REGION Network 65: SOLICITAÇÃO DE DESLIGAMENTO DO GRUPO 1
   RUNG wire#powerrail
      Contact( #AUX05 )
      wire#w1
      Contact( #LG1 )
      Contact( #G1L )
      Coil( #SDESG1 )
      wire#w2
      R_Coil( #LG1 )
   END_RUNG
   RUNG wire#powerrail
      Contact( #RTEOKG1 )
      Contact( #G1P )
   END_RUNG wire#w1
   RUNG wire#powerrail
      I_Contact( #G1OK )
   END_RUNG wire#w2
   RUNG wire#powerrail
      Contact( "AlwaysFALSE" )
      { S7_Templates := "SrcType := Int" } EQ_Contact(in1 := #NGS, in2 := 1)
      I_Contact( #G1P )
   END_RUNG wire#w2
   RUNG wire#powerrail
      Contact( "AlwaysFALSE" )
      { S7_Templates := "SrcType := Int" } EQ_Contact(in1 := #NGS, in2 := 2)
      I_Contact( #G1P )
      I_Contact( #G1C1 )
   END_RUNG wire#w2
   RUNG wire#powerrail
      Contact( "AlwaysFALSE" )
      { S7_Templates := "SrcType := Int" } EQ_Contact(in1 := #NGS, in2 := 3)
      I_Contact( #G1P )
      I_Contact( #G1C1 )
      I_Contact( #G1C2 )
   END_RUNG wire#w2
   RUNG wire#powerrail
      Contact( "AlwaysFALSE" )
      { S7_Templates := "SrcType := Int" } EQ_Contact(in1 := #NGS, in2 := 4)
      I_Contact( #G1P )
      I_Contact( #G1C1 )
      I_Contact( #G1C2 )
      I_Contact( #G1C3 )
   END_RUNG wire#w2
   // the same network as SCL:
   #SDESG1 := (#AUX05 OR (#RTEOKG1 AND #G1P)) AND #LG1 AND #G1L;
   IF #SDESG1 OR NOT #G1OK OR ("AlwaysFALSE" AND (#NGS = 1) AND NOT #G1P) OR ("AlwaysFALSE" AND (#NGS = 2) AND NOT #G1P AND NOT #G1C1) OR ("AlwaysFALSE" AND (#NGS = 3) AND NOT #G1P AND NOT #G1C1 AND NOT #G1C2) OR ("AlwaysFALSE" AND (#NGS = 4) AND NOT #G1P AND NOT #G1C1 AND NOT #G1C2 AND NOT #G1C3) THEN
       #LG1 := FALSE;
   END_IF;
END_REGION

REGION Network 66: SOLICITAÇÃO DE DESLIGAMENTO DO GRUPO 2
   #TSDG2(IN := (#SO_D OR NOT #DESAB) AND #G2P, PT := T#5S, ET => #ETTSDG2);   // TON
   #AUX06 := #TSDG2.Q;
END_REGION

REGION Network 67: SOLICITAÇÃO DE DESLIGAMENTO DO GRUPO 2
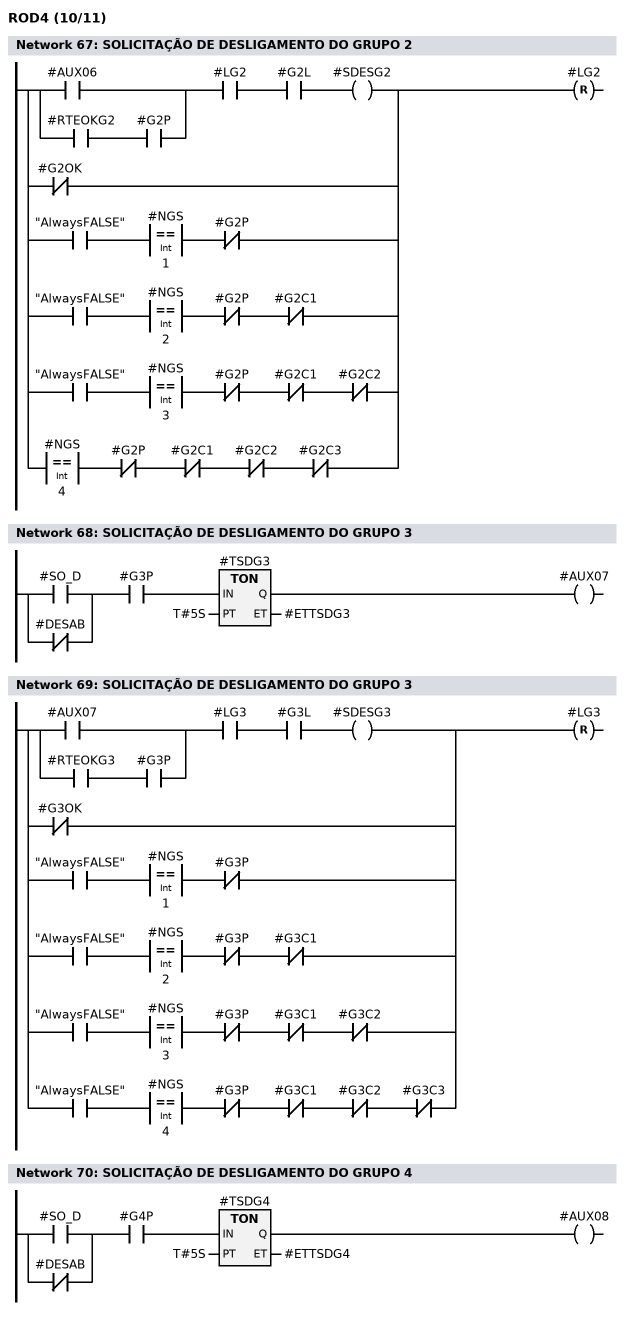
   RUNG wire#powerrail
      Contact( #AUX06 )
      wire#w1
      Contact( #LG2 )
      Contact( #G2L )
      Coil( #SDESG2 )
      wire#w2
      R_Coil( #LG2 )
   END_RUNG
   RUNG wire#powerrail
      Contact( #RTEOKG2 )
      Contact( #G2P )
   END_RUNG wire#w1
   RUNG wire#powerrail
      I_Contact( #G2OK )
   END_RUNG wire#w2
   RUNG wire#powerrail
      Contact( "AlwaysFALSE" )
      { S7_Templates := "SrcType := Int" } EQ_Contact(in1 := #NGS, in2 := 1)
      I_Contact( #G2P )
   END_RUNG wire#w2
   RUNG wire#powerrail
      Contact( "AlwaysFALSE" )
      { S7_Templates := "SrcType := Int" } EQ_Contact(in1 := #NGS, in2 := 2)
      I_Contact( #G2P )
      I_Contact( #G2C1 )
   END_RUNG wire#w2
   RUNG wire#powerrail
      Contact( "AlwaysFALSE" )
      { S7_Templates := "SrcType := Int" } EQ_Contact(in1 := #NGS, in2 := 3)
      I_Contact( #G2P )
      I_Contact( #G2C1 )
      I_Contact( #G2C2 )
   END_RUNG wire#w2
   RUNG wire#powerrail
      { S7_Templates := "SrcType := Int" } EQ_Contact(in1 := #NGS, in2 := 4)
      I_Contact( #G2P )
      I_Contact( #G2C1 )
      I_Contact( #G2C2 )
      I_Contact( #G2C3 )
   END_RUNG wire#w2
   // the same network as SCL:
   #SDESG2 := (#AUX06 OR (#RTEOKG2 AND #G2P)) AND #LG2 AND #G2L;
   IF #SDESG2 OR NOT #G2OK OR ("AlwaysFALSE" AND (#NGS = 1) AND NOT #G2P) OR ("AlwaysFALSE" AND (#NGS = 2) AND NOT #G2P AND NOT #G2C1) OR ("AlwaysFALSE" AND (#NGS = 3) AND NOT #G2P AND NOT #G2C1 AND NOT #G2C2) OR ((#NGS = 4) AND NOT #G2P AND NOT #G2C1 AND NOT #G2C2 AND NOT #G2C3) THEN
       #LG2 := FALSE;
   END_IF;
END_REGION

REGION Network 68: SOLICITAÇÃO DE DESLIGAMENTO DO GRUPO 3
   #TSDG3(IN := (#SO_D OR NOT #DESAB) AND #G3P, PT := T#5S, ET => #ETTSDG3);   // TON
   #AUX07 := #TSDG3.Q;
END_REGION

REGION Network 69: SOLICITAÇÃO DE DESLIGAMENTO DO GRUPO 3
   RUNG wire#powerrail
      Contact( #AUX07 )
      wire#w1
      Contact( #LG3 )
      Contact( #G3L )
      Coil( #SDESG3 )
      wire#w2
      R_Coil( #LG3 )
   END_RUNG
   RUNG wire#powerrail
      Contact( #RTEOKG3 )
      Contact( #G3P )
   END_RUNG wire#w1
   RUNG wire#powerrail
      I_Contact( #G3OK )
   END_RUNG wire#w2
   RUNG wire#powerrail
      Contact( "AlwaysFALSE" )
      { S7_Templates := "SrcType := Int" } EQ_Contact(in1 := #NGS, in2 := 1)
      I_Contact( #G3P )
   END_RUNG wire#w2
   RUNG wire#powerrail
      Contact( "AlwaysFALSE" )
      { S7_Templates := "SrcType := Int" } EQ_Contact(in1 := #NGS, in2 := 2)
      I_Contact( #G3P )
      I_Contact( #G3C1 )
   END_RUNG wire#w2
   RUNG wire#powerrail
      Contact( "AlwaysFALSE" )
      { S7_Templates := "SrcType := Int" } EQ_Contact(in1 := #NGS, in2 := 3)
      I_Contact( #G3P )
      I_Contact( #G3C1 )
      I_Contact( #G3C2 )
   END_RUNG wire#w2
   RUNG wire#powerrail
      Contact( "AlwaysFALSE" )
      { S7_Templates := "SrcType := Int" } EQ_Contact(in1 := #NGS, in2 := 4)
      I_Contact( #G3P )
      I_Contact( #G3C1 )
      I_Contact( #G3C2 )
      I_Contact( #G3C3 )
   END_RUNG wire#w2
   // the same network as SCL:
   #SDESG3 := (#AUX07 OR (#RTEOKG3 AND #G3P)) AND #LG3 AND #G3L;
   IF #SDESG3 OR NOT #G3OK OR ("AlwaysFALSE" AND (#NGS = 1) AND NOT #G3P) OR ("AlwaysFALSE" AND (#NGS = 2) AND NOT #G3P AND NOT #G3C1) OR ("AlwaysFALSE" AND (#NGS = 3) AND NOT #G3P AND NOT #G3C1 AND NOT #G3C2) OR ("AlwaysFALSE" AND (#NGS = 4) AND NOT #G3P AND NOT #G3C1 AND NOT #G3C2 AND NOT #G3C3) THEN
       #LG3 := FALSE;
   END_IF;
END_REGION

REGION Network 70: SOLICITAÇÃO DE DESLIGAMENTO DO GRUPO 4
   #TSDG4(IN := (#SO_D OR NOT #DESAB) AND #G4P, PT := T#5S, ET => #ETTSDG4);   // TON
   #AUX08 := #TSDG4.Q;
END_REGION

REGION Network 71: SOLICITAÇÃO DE DESLIGAMENTO DO GRUPO 4
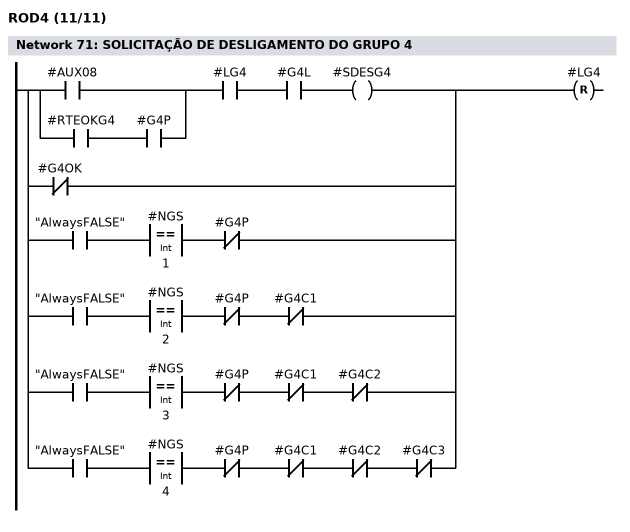
   RUNG wire#powerrail
      Contact( #AUX08 )
      wire#w1
      Contact( #LG4 )
      Contact( #G4L )
      Coil( #SDESG4 )
      wire#w2
      R_Coil( #LG4 )
   END_RUNG
   RUNG wire#powerrail
      Contact( #RTEOKG4 )
      Contact( #G4P )
   END_RUNG wire#w1
   RUNG wire#powerrail
      I_Contact( #G4OK )
   END_RUNG wire#w2
   RUNG wire#powerrail
      Contact( "AlwaysFALSE" )
      { S7_Templates := "SrcType := Int" } EQ_Contact(in1 := #NGS, in2 := 1)
      I_Contact( #G4P )
   END_RUNG wire#w2
   RUNG wire#powerrail
      Contact( "AlwaysFALSE" )
      { S7_Templates := "SrcType := Int" } EQ_Contact(in1 := #NGS, in2 := 2)
      I_Contact( #G4P )
      I_Contact( #G4C1 )
   END_RUNG wire#w2
   RUNG wire#powerrail
      Contact( "AlwaysFALSE" )
      { S7_Templates := "SrcType := Int" } EQ_Contact(in1 := #NGS, in2 := 3)
      I_Contact( #G4P )
      I_Contact( #G4C1 )
      I_Contact( #G4C2 )
   END_RUNG wire#w2
   RUNG wire#powerrail
      Contact( "AlwaysFALSE" )
      { S7_Templates := "SrcType := Int" } EQ_Contact(in1 := #NGS, in2 := 4)
      I_Contact( #G4P )
      I_Contact( #G4C1 )
      I_Contact( #G4C2 )
      I_Contact( #G4C3 )
   END_RUNG wire#w2
   // the same network as SCL:
   #SDESG4 := (#AUX08 OR (#RTEOKG4 AND #G4P)) AND #LG4 AND #G4L;
   IF #SDESG4 OR NOT #G4OK OR ("AlwaysFALSE" AND (#NGS = 1) AND NOT #G4P) OR ("AlwaysFALSE" AND (#NGS = 2) AND NOT #G4P AND NOT #G4C1) OR ("AlwaysFALSE" AND (#NGS = 3) AND NOT #G4P AND NOT #G4C1 AND NOT #G4C2) OR ("AlwaysFALSE" AND (#NGS = 4) AND NOT #G4P AND NOT #G4C1 AND NOT #G4C2 AND NOT #G4C3) THEN
       #LG4 := FALSE;
   END_IF;
END_REGION
END_FUNCTION_BLOCK

FUNCTION_BLOCK "INSTRUMENTO"   // FB201, LAD
TITLE = BLOCO PARA CONVERSÃO DE ESCALA DE ENGENHARIA
{ S7_Optimized_Access := 'FALSE' }
VERSION : 0.1
   VAR_INPUT
      "VALOR MANUAL" : Real;   // VALOR MANUAL (HMI)
      EA : Int;   // LEITURA DO CANAL ANALÓGICO
      EA_IE : Real;   // INÍCIO DA ESCALA DO CANAL
      EA_FE : Real;   // FIM DE ESCALA DO CANAL
      S_IE : Real;   // INÍCIO DE ESCALA DE ENGENHARIA PRINCIPAL
      S_FE : Real;   // FIM DE ESCALA DE ENGENHARIA PRINCIPAL
      S2_IE : Real;   // INÍCIO DE ESCALA DE ENGENHARIA SECUNDÁRIA
      S2_FE : Real;   // FIM DE ESCALA DE ENGENHARIA SECUNDÁRIA
      SPLL : Real;   // SETPOINT MUITO BAIXO
      SPL : Real;   // SETPOINT BAIXO
      SPH : Real;   // SETPOINT ALTO
      SPHH : Real;   // SETPOINT MUITO ALTO
      TE_LL : Time;   // DELAY PARA ALARME MUITO BAIXO
      TE_L : Time;   // DELAY PARA ALARME BAIXO
      TE_H : Time;   // DELAY PARA ALARME ALTO
      TE_HH : Time;   // DELAY PARA ALARME MUITO ALTO
      FRH : Int;   // VALOR ALTO PARA ALARME DE FALHA DE LEITURA
      FRL : Int;   // VALOR BAIXO PARA ALARME DE FALHA DE LEITURA
      LIM : Bool;   // LIMITA O VALOR À ESCALA
      MANUAL : Bool;   // HABILITA MANUTENÇÃO DO INSTRUMENTO
      COND : Bool;   // CONDIÇÃO PARA GERAR ALARME
      SPR_YLL : Bool;   // HABILITA SUPRESSÃO ALARME MUITO BAIXO
      SPR_YL : Bool;   // HABILITA SUPRESSÃO ALARME BAIXO
      SPR_YH : Bool;   // HABILITA SUPRESSÃO ALARME ALTO
      SPR_YHH : Bool;   // HABILITA SUPRESSÃO ALARME MUITO ALTO
   END_VAR
   VAR_OUTPUT
      VNP : Real;   // VALOR CONVERTIDO PARA ESCALA DE ENGENHARIA PRINCIPAL
      YLL : Bool;   // ALARME MUITO BAIXO
      YL : Bool;   // ALARME BAIXO
      YH : Bool;   // ALARME ALTO
      YHH : Bool;   // ALARME MUITO ALTO
      YF : Bool;   // ALARME DE FALHA NA MEDIÇÃO
      VNS : Real;   // VALOR CONVERTIDO PARA ESCALA DE ENGENHARIA SECUNDÁRIA
      LL : Bool;   // VALOR MUITO BAIXO
      L : Bool;   // VALOR BAIXO
      H : Bool;   // VALOR ALTO
      HH : Bool;   // VALOR MUITO ALTO
   END_VAR
   VAR
      TLL : TON_TIME;   // TEMPO PARA GERAR ALARME
      TL : TON_TIME;   // TEMPO PARA GERAR ALARME
      TH : TON_TIME;   // TEMPO PARA GERAR ALARME
      THH : TON_TIME;   // TEMPO PARA GERAR ALARME
      FALHA : Bool;   // SINALIZAÇÃO DE FALHA NO INSTRUMENTO
   END_VAR
   VAR_TEMP
      EAR : Real;   // VALOR LIDO DA ENTRADA ANALÓGICA
      AC01 : Real;   // AUXILIAR PARA CÁLCULO
      AC02 : Real;   // AUXILIAR PARA CÁLCULO
      AC03 : Real;   // AUXILIAR PARA CÁLCULO
      AC04 : Real;   // AUXILIAR PARA CÁLCULO
      AC05 : Real;   // AUXILIAR PARA CÁLCULO
      AC06 : Real;   // AUXILIAR PARA CÁLCULO
      AC07 : Real;   // AUXILIAR PARA CÁLCULO
      AC08 : Real;   // AUXILIAR PARA CÁLCULO
      AC09 : Real;   // AUXILIAR PARA CÁLCULO
      AC10 : Real;   // AUXILIAR PARA CÁLCULO
      RESULT_P : Real;   // RESULTADO DA ESCALA
      RESULT_S : Real;   // RESULTADO DA ESCALA
      ET_TLL : Time;   // EFETIVO DO TEMPORIZADOR
      ET_TL : Time;   // EFETIVO DO TEMPORIZADOR
      ET_TH : Time;   // EFETIVO DO TEMPORIZADOR
      ET_THH : Time;   // EFETIVO DO TEMPORIZADOR
      EADI : DInt;
   END_VAR
BEGIN

REGION Network 1: CONVERSOR O VALOR LIDO DO CARTÃO PARA REAL
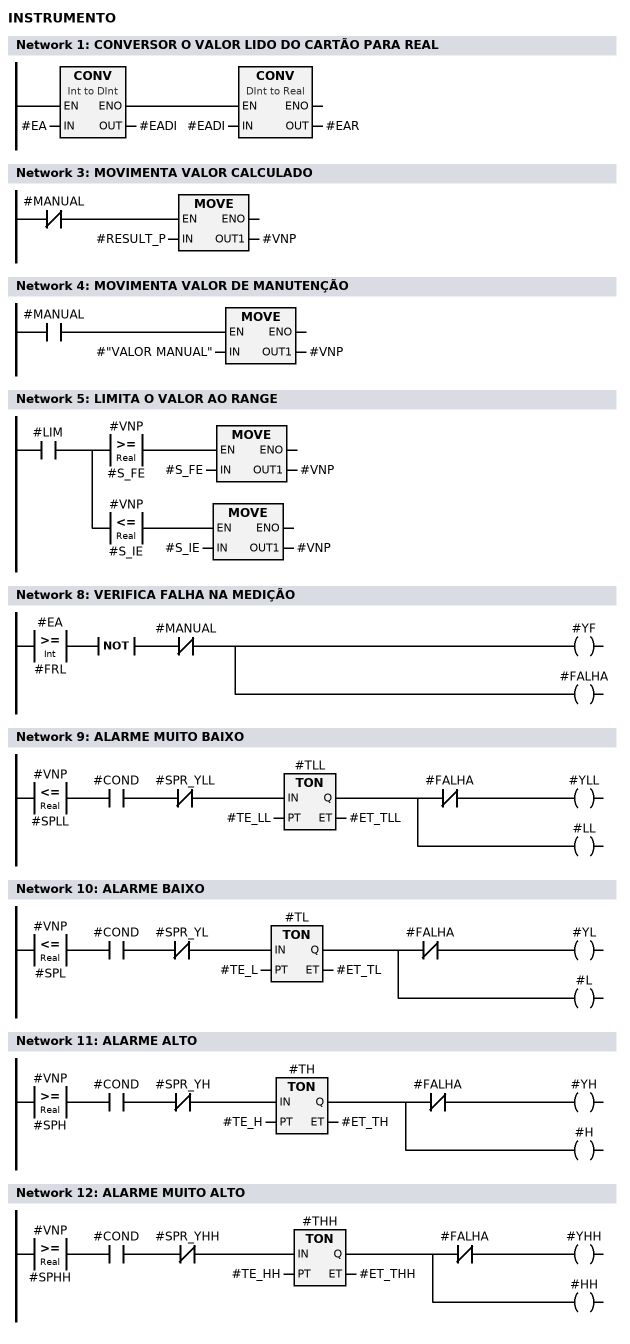
   RUNG wire#powerrail
      { S7_Templates := "[SrcType := Int, DestType := DInt]"; S7_GenerateENO := "TRUE" } Convert(in := #EA, out => #EADI)
      { S7_Templates := "[SrcType := DInt, DestType := Real]"; S7_GenerateENO := "TRUE" } Convert(in := #EADI, out => #EAR)
   END_RUNG
   // the same network as SCL:
   // ENO of a box is taken as its EN; it also drops when the box reports an error
   #EADI := INT_TO_DINT(#EA);
   #EAR := DINT_TO_REAL(#EADI);
END_REGION

REGION Network 2 (STL): CONVERTER PARA ESCALA DE ENGENHARIA PRINCIPAL
         L     #EAR;
         L     #EA_IE;
         -R;
         T     #AC01;

         L     #S_FE;  // Subtrai escalas de saída
         L     #S_IE;
         -R;
         T     #AC02;

         L     #EA_FE;  // Subtrai escalas de entrada
         L     #EA_IE;
         -R;
         T     #AC03;

         L     #AC01;  // Multiplica resultado das subtrações
         L     #AC02;
         *R;
         T     #AC04;

         L     #AC04;  // Divide o produto pela subtração das escalas de entrada
         L     #AC03;
         /R;
         T     #AC05;

         L     #AC05;  // Soma o valor de fim da escala de saída
         L     #S_IE;
         +R;
         T     #RESULT_P;  // Resultado do cálculo
         T     #VNP;  // Transfere valor já convertido
END_REGION

REGION Network 3: MOVIMENTA VALOR CALCULADO
   RUNG wire#powerrail
      I_Contact( #MANUAL )
      Move(in := #RESULT_P, out1 => #VNP)
   END_RUNG
   // the same network as SCL:
   IF NOT #MANUAL THEN #VNP := #RESULT_P; END_IF;
END_REGION

REGION Network 4: MOVIMENTA VALOR DE MANUTENÇÃO
   RUNG wire#powerrail
      Contact( #MANUAL )
      Move(in := #"VALOR MANUAL", out1 => #VNP)
   END_RUNG
   // the same network as SCL:
   IF #MANUAL THEN #VNP := #"VALOR MANUAL"; END_IF;
END_REGION

REGION Network 5: LIMITA O VALOR AO RANGE
   RUNG wire#powerrail
      Contact( #LIM )
      wire#w1
      { S7_Templates := "SrcType := Real" } GE_Contact(in1 := #VNP, in2 := #S_FE)
      { S7_GenerateENO := "TRUE" } Move(in := #S_FE, out1 => #VNP)
   END_RUNG
   RUNG wire#w1
      { S7_Templates := "SrcType := Real" } LE_Contact(in1 := #VNP, in2 := #S_IE)
      { S7_GenerateENO := "TRUE" } Move(in := #S_IE, out1 => #VNP)
   END_RUNG
   // the same network as SCL:
   IF #LIM AND (#VNP >= #S_FE) THEN #VNP := #S_FE; END_IF;
   IF #LIM AND (#VNP <= #S_IE) THEN #VNP := #S_IE; END_IF;
END_REGION

REGION Network 6 (STL): MOVIMENTA 0 PARA A LEITURA
         A     #YF;
         AN    #MANUAL;
         JNB   _004;
         L     0;
         T     #VNP;
   _004: NOP   0;
END_REGION

REGION Network 7 (STL): CONVERTER PARA ESCALA DE ENGENHARIA SECUNDÁRIA
         L     #VNP;
         L     #S_IE;
         -R;
         T     #AC06;

         L     #S2_FE;  // Subtrai escalas de saída
         L     #S2_IE;
         -R;
         T     #AC07;

         L     #S_FE;  // Subtrai escalas de entrada
         L     #S_IE;
         -R;
         T     #AC08;

         L     #AC06;  // Multiplica resultado das subtrações
         L     #AC07;
         *R;
         T     #AC09;

         L     #AC09;  // Divide o produto pela subtração das escalas de entrada
         L     #AC08;
         /R;
         T     #AC10;

         L     #AC10;  // Soma o valor de fim da escala de saída
         L     #S2_IE;
         +R;
         T     #RESULT_S;  // Resultado do cálculo
         T     #VNS;  // Transfere valor já convertido
END_REGION

REGION Network 8: VERIFICA FALHA NA MEDIÇÃO
   RUNG wire#powerrail
      { S7_Templates := "SrcType := Int" } GE_Contact(in1 := #EA, in2 := #FRL)
      Not()
      I_Contact( #MANUAL )
      wire#w1
      Coil( #YF )
   END_RUNG
   RUNG wire#w1
      Coil( #FALHA )
   END_RUNG
   // the same network as SCL:
   #YF := NOT (#EA >= #FRL) AND NOT #MANUAL;
   #FALHA := #YF;
END_REGION

REGION Network 9: ALARME MUITO BAIXO
   #TLL(IN := (#VNP <= #SPLL) AND #COND AND NOT #SPR_YLL, PT := #TE_LL, ET => #ET_TLL);   // TON
   #YLL := #TLL.Q AND NOT #FALHA;
   #LL := #TLL.Q;
END_REGION

REGION Network 10: ALARME BAIXO
   #TL(IN := (#VNP <= #SPL) AND #COND AND NOT #SPR_YL, PT := #TE_L, ET => #ET_TL);   // TON
   #YL := #TL.Q AND NOT #FALHA;
   #L := #TL.Q;
END_REGION

REGION Network 11: ALARME ALTO
   #TH(IN := (#VNP >= #SPH) AND #COND AND NOT #SPR_YH, PT := #TE_H, ET => #ET_TH);   // TON
   #YH := #TH.Q AND NOT #FALHA;
   #H := #TH.Q;
END_REGION

REGION Network 12: ALARME MUITO ALTO
   #THH(IN := (#VNP >= #SPHH) AND #COND AND NOT #SPR_YHH, PT := #TE_HH, ET => #ET_THH);   // TON
   #YHH := #THH.Q AND NOT #FALHA;
   #HH := #THH.Q;
END_REGION
END_FUNCTION_BLOCK

FUNCTION_BLOCK "INTPRO"   // FB202, LAD
{ S7_Optimized_Access := 'FALSE' }
VERSION : 0.1
   VAR
      EE_P_NIV : Bool;   // HAILITA BOMBA PRINCIPAL PELO NÍVEL
      EE_C1_NIV : Bool;   // HAILITA BOMBA COMPLEMENTAR 1 PELO NÍVEL
      EE_C2_NIV : Bool;   // HAILITA BOMBA COMPLEMENTAR 2 PELO NÍVEL
      EE_P_LS : Bool;   // HAILITA BOMBA PRINCIPAL PELAS BÓIAS
      EE_C1_LS : Bool;   // HAILITA BOMBA COMLEMENTAR 1 PELAS BÓIAS
      EE_C2_LS : Bool;   // HAILITA BOMBA COMPLEMENTAR 2 PELAS BÓIAS
      HAB_P_EE : Bool;   // LIGA BOMBA PRINCIPAL DA ELEVATÓRIA
      HAB_C1_EE : Bool;   // LIGA BOMBA COMPLEMENTAR 1 DA ELEVATÓRIA
      HAB_C2_EE : Bool;   // LIGA BOMBA COMPLEMENTAR 2 DA ELEVATÓRIA
      AUXP01 : Bool;
      BS01OK : Bool;
      BS02OK : Bool;
      BS03OK : Bool;
      L_BS01 : Bool;
      L_BS02 : Bool;
      L_BS03 : Bool;
      AUXP02 : Bool;
      AUXP03 : Bool;
      AUXP04 : Bool;
      AUXP05 : Bool;
      AUXP06 : Bool;
      AUXP07 : Bool;
      ETBS01_T001 : Int;
      ETBS02_T001 : Int;
      ETBS03_T001 : Int;
      BS01TO : Int;
      BS02TO : Int;
      BS03TO : Int;
      BS01TEOK : DInt;
      BS02TEOK : DInt;
      BS03TEOK : DInt;
      TE00 : IEC_TIMER;
      RODEE : "ROD4";
   END_VAR
   VAR_TEMP
      T011S : Int;
      ET_TE00 : Time;
   END_VAR
BEGIN

REGION Network 1: Alarme falha de sinal transmissor de nivel
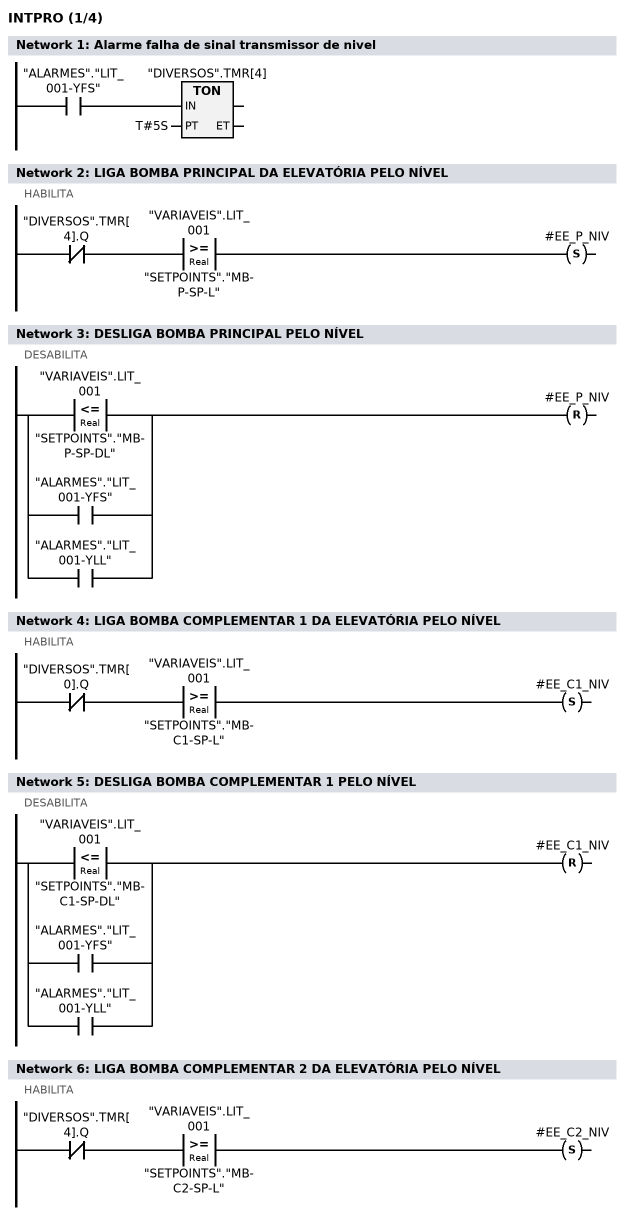
   "DIVERSOS".TMR[4].TON(IN := "ALARMES"."LIT_001-YFS", PT := T#5S);
END_REGION

REGION Network 2: LIGA BOMBA PRINCIPAL DA ELEVATÓRIA PELO NÍVEL
   // HABILITA
   RUNG wire#powerrail
      I_Contact( "DIVERSOS".TMR[4].Q )
      { S7_Templates := "SrcType := Real" } GE_Contact(in1 := "VARIAVEIS".LIT_001, in2 := "SETPOINTS"."MB-P-SP-L")
      S_Coil( #EE_P_NIV )
   END_RUNG
   // the same network as SCL:
   IF NOT "DIVERSOS".TMR[4].Q AND ("VARIAVEIS".LIT_001 >= "SETPOINTS"."MB-P-SP-L") THEN
       #EE_P_NIV := TRUE;
   END_IF;
END_REGION

REGION Network 3: DESLIGA BOMBA PRINCIPAL PELO NÍVEL
   // DESABILITA
   RUNG wire#powerrail
      { S7_Templates := "SrcType := Real" } LE_Contact(in1 := "VARIAVEIS".LIT_001, in2 := "SETPOINTS"."MB-P-SP-DL")
      wire#w1
      R_Coil( #EE_P_NIV )
   END_RUNG
   RUNG wire#powerrail
      Contact( "ALARMES"."LIT_001-YFS" )
   END_RUNG wire#w1
   RUNG wire#powerrail
      Contact( "ALARMES"."LIT_001-YLL" )
   END_RUNG wire#w1
   // the same network as SCL:
   IF ("VARIAVEIS".LIT_001 <= "SETPOINTS"."MB-P-SP-DL") OR "ALARMES"."LIT_001-YFS" OR "ALARMES"."LIT_001-YLL" THEN
       #EE_P_NIV := FALSE;
   END_IF;
END_REGION

REGION Network 4: LIGA BOMBA COMPLEMENTAR 1 DA ELEVATÓRIA PELO NÍVEL
   // HABILITA
   RUNG wire#powerrail
      I_Contact( "DIVERSOS".TMR[0].Q )
      { S7_Templates := "SrcType := Real" } GE_Contact(in1 := "VARIAVEIS".LIT_001, in2 := "SETPOINTS"."MB-C1-SP-L")
      S_Coil( #EE_C1_NIV )
   END_RUNG
   // the same network as SCL:
   IF NOT "DIVERSOS".TMR[0].Q AND ("VARIAVEIS".LIT_001 >= "SETPOINTS"."MB-C1-SP-L") THEN
       #EE_C1_NIV := TRUE;
   END_IF;
END_REGION

REGION Network 5: DESLIGA BOMBA COMPLEMENTAR 1 PELO NÍVEL
   // DESABILITA
   RUNG wire#powerrail
      { S7_Templates := "SrcType := Real" } LE_Contact(in1 := "VARIAVEIS".LIT_001, in2 := "SETPOINTS"."MB-C1-SP-DL")
      wire#w1
      R_Coil( #EE_C1_NIV )
   END_RUNG
   RUNG wire#powerrail
      Contact( "ALARMES"."LIT_001-YFS" )
   END_RUNG wire#w1
   RUNG wire#powerrail
      Contact( "ALARMES"."LIT_001-YLL" )
   END_RUNG wire#w1
   // the same network as SCL:
   IF ("VARIAVEIS".LIT_001 <= "SETPOINTS"."MB-C1-SP-DL") OR "ALARMES"."LIT_001-YFS" OR "ALARMES"."LIT_001-YLL" THEN
       #EE_C1_NIV := FALSE;
   END_IF;
END_REGION

REGION Network 6: LIGA BOMBA COMPLEMENTAR 2 DA ELEVATÓRIA PELO NÍVEL
   // HABILITA
   RUNG wire#powerrail
      I_Contact( "DIVERSOS".TMR[4].Q )
      { S7_Templates := "SrcType := Real" } GE_Contact(in1 := "VARIAVEIS".LIT_001, in2 := "SETPOINTS"."MB-C2-SP-L")
      S_Coil( #EE_C2_NIV )
   END_RUNG
   // the same network as SCL:
   IF NOT "DIVERSOS".TMR[4].Q AND ("VARIAVEIS".LIT_001 >= "SETPOINTS"."MB-C2-SP-L") THEN
       #EE_C2_NIV := TRUE;
   END_IF;
END_REGION

REGION Network 7: DESLIGA BOMBA COMPLEMENTAR 2 PELO NÍVEL
   // DESABILITA
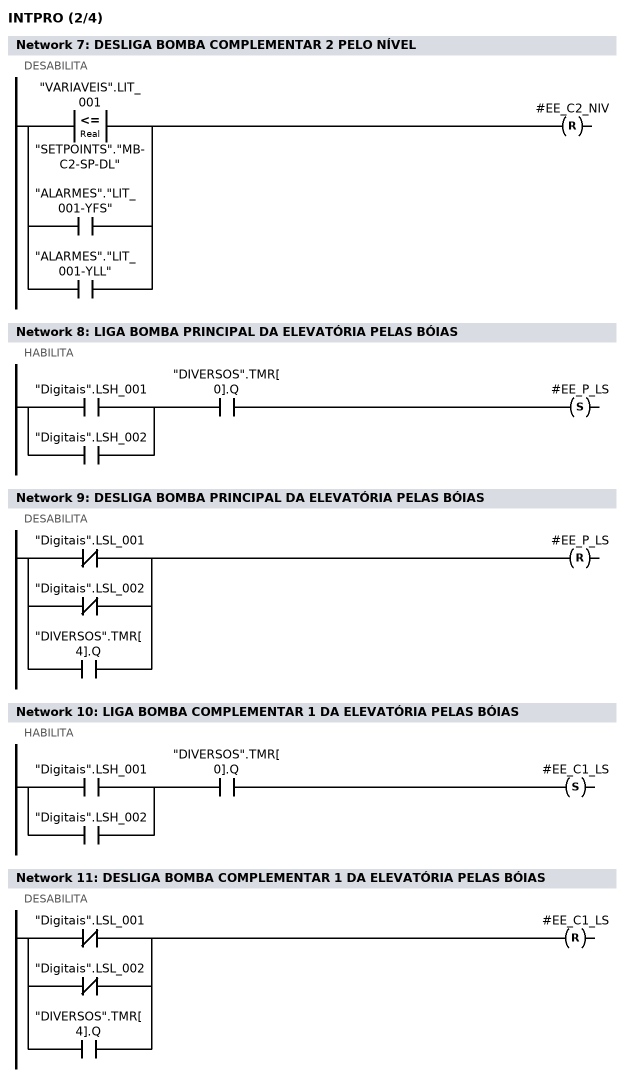
   RUNG wire#powerrail
      { S7_Templates := "SrcType := Real" } LE_Contact(in1 := "VARIAVEIS".LIT_001, in2 := "SETPOINTS"."MB-C2-SP-DL")
      wire#w1
      R_Coil( #EE_C2_NIV )
   END_RUNG
   RUNG wire#powerrail
      Contact( "ALARMES"."LIT_001-YFS" )
   END_RUNG wire#w1
   RUNG wire#powerrail
      Contact( "ALARMES"."LIT_001-YLL" )
   END_RUNG wire#w1
   // the same network as SCL:
   IF ("VARIAVEIS".LIT_001 <= "SETPOINTS"."MB-C2-SP-DL") OR "ALARMES"."LIT_001-YFS" OR "ALARMES"."LIT_001-YLL" THEN
       #EE_C2_NIV := FALSE;
   END_IF;
END_REGION

REGION Network 8: LIGA BOMBA PRINCIPAL DA ELEVATÓRIA PELAS BÓIAS
   // HABILITA
   RUNG wire#powerrail
      Contact( "Digitais".LSH_001 )
      wire#w1
      Contact( "DIVERSOS".TMR[0].Q )
      S_Coil( #EE_P_LS )
   END_RUNG
   RUNG wire#powerrail
      Contact( "Digitais".LSH_002 )
   END_RUNG wire#w1
   // the same network as SCL:
   IF ("Digitais".LSH_001 OR "Digitais".LSH_002) AND "DIVERSOS".TMR[0].Q THEN #EE_P_LS := TRUE; END_IF;
END_REGION

REGION Network 9: DESLIGA BOMBA PRINCIPAL DA ELEVATÓRIA PELAS BÓIAS
   // DESABILITA
   RUNG wire#powerrail
      I_Contact( "Digitais".LSL_001 )
      wire#w1
      R_Coil( #EE_P_LS )
   END_RUNG
   RUNG wire#powerrail
      I_Contact( "Digitais".LSL_002 )
   END_RUNG wire#w1
   RUNG wire#powerrail
      Contact( "DIVERSOS".TMR[4].Q )
   END_RUNG wire#w1
   // the same network as SCL:
   IF NOT "Digitais".LSL_001 OR NOT "Digitais".LSL_002 OR "DIVERSOS".TMR[4].Q THEN #EE_P_LS := FALSE; END_IF;
END_REGION

REGION Network 10: LIGA BOMBA COMPLEMENTAR 1 DA ELEVATÓRIA PELAS BÓIAS
   // HABILITA
   RUNG wire#powerrail
      Contact( "Digitais".LSH_001 )
      wire#w1
      Contact( "DIVERSOS".TMR[0].Q )
      S_Coil( #EE_C1_LS )
   END_RUNG
   RUNG wire#powerrail
      Contact( "Digitais".LSH_002 )
   END_RUNG wire#w1
   // the same network as SCL:
   IF ("Digitais".LSH_001 OR "Digitais".LSH_002) AND "DIVERSOS".TMR[0].Q THEN #EE_C1_LS := TRUE; END_IF;
END_REGION

REGION Network 11: DESLIGA BOMBA COMPLEMENTAR 1 DA ELEVATÓRIA PELAS BÓIAS
   // DESABILITA
   RUNG wire#powerrail
      I_Contact( "Digitais".LSL_001 )
      wire#w1
      R_Coil( #EE_C1_LS )
   END_RUNG
   RUNG wire#powerrail
      I_Contact( "Digitais".LSL_002 )
   END_RUNG wire#w1
   RUNG wire#powerrail
      Contact( "DIVERSOS".TMR[4].Q )
   END_RUNG wire#w1
   // the same network as SCL:
   IF NOT "Digitais".LSL_001 OR NOT "Digitais".LSL_002 OR "DIVERSOS".TMR[4].Q THEN
       #EE_C1_LS := FALSE;
   END_IF;
END_REGION

REGION Network 12: LIGA BOMBA COMPLEMENTAR 2 DA ELEVATÓRIA PELAS BÓIAS
   // HABILITA
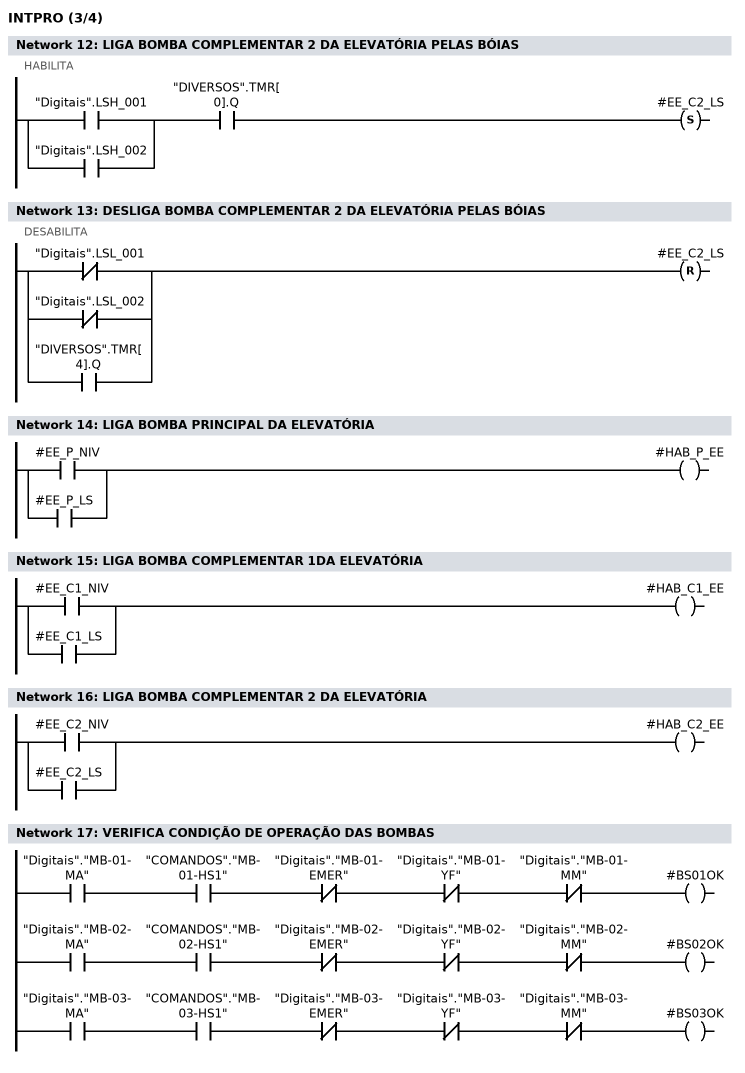
   RUNG wire#powerrail
      Contact( "Digitais".LSH_001 )
      wire#w1
      Contact( "DIVERSOS".TMR[0].Q )
      S_Coil( #EE_C2_LS )
   END_RUNG
   RUNG wire#powerrail
      Contact( "Digitais".LSH_002 )
   END_RUNG wire#w1
   // the same network as SCL:
   IF ("Digitais".LSH_001 OR "Digitais".LSH_002) AND "DIVERSOS".TMR[0].Q THEN #EE_C2_LS := TRUE; END_IF;
END_REGION

REGION Network 13: DESLIGA BOMBA COMPLEMENTAR 2 DA ELEVATÓRIA PELAS BÓIAS
   // DESABILITA
   RUNG wire#powerrail
      I_Contact( "Digitais".LSL_001 )
      wire#w1
      R_Coil( #EE_C2_LS )
   END_RUNG
   RUNG wire#powerrail
      I_Contact( "Digitais".LSL_002 )
   END_RUNG wire#w1
   RUNG wire#powerrail
      Contact( "DIVERSOS".TMR[4].Q )
   END_RUNG wire#w1
   // the same network as SCL:
   IF NOT "Digitais".LSL_001 OR NOT "Digitais".LSL_002 OR "DIVERSOS".TMR[4].Q THEN
       #EE_C2_LS := FALSE;
   END_IF;
END_REGION

REGION Network 14: LIGA BOMBA PRINCIPAL DA ELEVATÓRIA
   RUNG wire#powerrail
      Contact( #EE_P_NIV )
      wire#w1
      Coil( #HAB_P_EE )
   END_RUNG
   RUNG wire#powerrail
      Contact( #EE_P_LS )
   END_RUNG wire#w1
   // the same network as SCL:
   #HAB_P_EE := #EE_P_NIV OR #EE_P_LS;
END_REGION

REGION Network 15: LIGA BOMBA COMPLEMENTAR 1DA ELEVATÓRIA
   RUNG wire#powerrail
      Contact( #EE_C1_NIV )
      wire#w1
      Coil( #HAB_C1_EE )
   END_RUNG
   RUNG wire#powerrail
      Contact( #EE_C1_LS )
   END_RUNG wire#w1
   // the same network as SCL:
   #HAB_C1_EE := #EE_C1_NIV OR #EE_C1_LS;
END_REGION

REGION Network 16: LIGA BOMBA COMPLEMENTAR 2 DA ELEVATÓRIA
   RUNG wire#powerrail
      Contact( #EE_C2_NIV )
      wire#w1
      Coil( #HAB_C2_EE )
   END_RUNG
   RUNG wire#powerrail
      Contact( #EE_C2_LS )
   END_RUNG wire#w1
   // the same network as SCL:
   #HAB_C2_EE := #EE_C2_NIV OR #EE_C2_LS;
END_REGION

REGION Network 17: VERIFICA CONDIÇÃO DE OPERAÇÃO DAS BOMBAS
   RUNG wire#powerrail
      Contact( "Digitais"."MB-01-MA" )
      Contact( "COMANDOS"."MB-01-HS1" )
      I_Contact( "Digitais"."MB-01-EMER" )
      I_Contact( "Digitais"."MB-01-YF" )
      I_Contact( "Digitais"."MB-01-MM" )
      Coil( #BS01OK )
   END_RUNG
   RUNG wire#powerrail
      Contact( "Digitais"."MB-02-MA" )
      Contact( "COMANDOS"."MB-02-HS1" )
      I_Contact( "Digitais"."MB-02-EMER" )
      I_Contact( "Digitais"."MB-02-YF" )
      I_Contact( "Digitais"."MB-02-MM" )
      Coil( #BS02OK )
   END_RUNG
   RUNG wire#powerrail
      Contact( "Digitais"."MB-03-MA" )
      Contact( "COMANDOS"."MB-03-HS1" )
      I_Contact( "Digitais"."MB-03-EMER" )
      I_Contact( "Digitais"."MB-03-YF" )
      I_Contact( "Digitais"."MB-03-MM" )
      Coil( #BS03OK )
   END_RUNG
   // the same network as SCL:
   #BS01OK := "Digitais"."MB-01-MA" AND "COMANDOS"."MB-01-HS1" AND NOT "Digitais"."MB-01-EMER" AND NOT "Digitais"."MB-01-YF" AND NOT "Digitais"."MB-01-MM";
   #BS02OK := "Digitais"."MB-02-MA" AND "COMANDOS"."MB-02-HS1" AND NOT "Digitais"."MB-02-EMER" AND NOT "Digitais"."MB-02-YF" AND NOT "Digitais"."MB-02-MM";
   #BS03OK := "Digitais"."MB-03-MA" AND "COMANDOS"."MB-03-HS1" AND NOT "Digitais"."MB-03-EMER" AND NOT "Digitais"."MB-03-YF" AND NOT "Digitais"."MB-03-MM";
END_REGION

REGION Network 18: RODÍZIO DAS BOMBAS
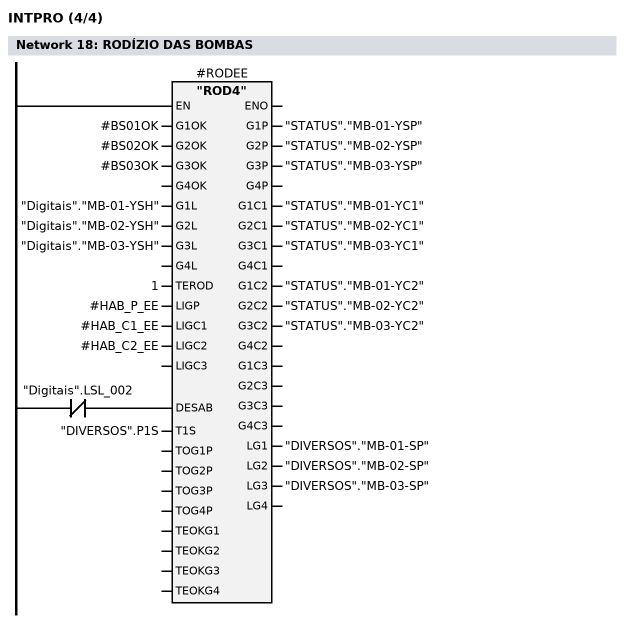
   RUNG wire#powerrail
      #RODEE(DESAB := wire#w1, G1OK := #BS01OK, G2OK := #BS02OK, G3OK := #BS03OK, G4OK :=, G1L := "Digitais"."MB-01-YSH", G2L := "Digitais"."MB-02-YSH", G3L := "Digitais"."MB-03-YSH", G4L :=, TEROD := 1, LIGP := #HAB_P_EE, LIGC1 := #HAB_C1_EE, LIGC2 := #HAB_C2_EE, LIGC3 :=, T1S := "DIVERSOS".P1S, TOG1P :=, TOG2P :=, TOG3P :=, TOG4P :=, TEOKG1 :=, TEOKG2 :=, TEOKG3 :=, TEOKG4 :=, G1P => "STATUS"."MB-01-YSP", G2P => "STATUS"."MB-02-YSP", G3P => "STATUS"."MB-03-YSP", G4P =>, G1C1 => "STATUS"."MB-01-YC1", G2C1 => "STATUS"."MB-02-YC1", G3C1 => "STATUS"."MB-03-YC1", G4C1 =>, G1C2 => "STATUS"."MB-01-YC2", G2C2 => "STATUS"."MB-02-YC2", G3C2 => "STATUS"."MB-03-YC2", G4C2 =>, G1C3 =>, G2C3 =>, G3C3 =>, G4C3 =>, LG1 => "DIVERSOS"."MB-01-SP", LG2 => "DIVERSOS"."MB-02-SP", LG3 => "DIVERSOS"."MB-03-SP", LG4 =>)
   END_RUNG
   RUNG wire#powerrail
      I_Contact( "Digitais".LSL_002 )
   END_RUNG wire#w1
   // the same network as SCL:
   #RODEE(G1OK := #BS01OK,   // "ROD4"
          G2OK := #BS02OK,
          G3OK := #BS03OK,
          G1L := "Digitais"."MB-01-YSH",
          G2L := "Digitais"."MB-02-YSH",
          G3L := "Digitais"."MB-03-YSH",
          TEROD := 1,
          LIGP := #HAB_P_EE,
          LIGC1 := #HAB_C1_EE,
          LIGC2 := #HAB_C2_EE,
          DESAB := NOT "Digitais".LSL_002,
          T1S := "DIVERSOS".P1S,
          G1P => "STATUS"."MB-01-YSP",
          G2P => "STATUS"."MB-02-YSP",
          G3P => "STATUS"."MB-03-YSP",
          G1C1 => "STATUS"."MB-01-YC1",
          G2C1 => "STATUS"."MB-02-YC1",
          G3C1 => "STATUS"."MB-03-YC1",
          G1C2 => "STATUS"."MB-01-YC2",
          G2C2 => "STATUS"."MB-02-YC2",
          G3C2 => "STATUS"."MB-03-YC2",
          LG1 => "DIVERSOS"."MB-01-SP",
          LG2 => "DIVERSOS"."MB-02-SP",
          LG3 => "DIVERSOS"."MB-03-SP");
END_REGION
END_FUNCTION_BLOCK

FUNCTION_BLOCK "ROD2"   // FB205, LAD
TITLE = RODÍZIO DE 2 GRUPOS
{ S7_Optimized_Access := 'FALSE' }
VERSION : 0.1
   VAR_INPUT
      G1OK : Bool;   // GRUPO EM CONDIÇÕES DE OPERAÇÃO
      G2OK : Bool;   // GRUPO EM CONDIÇÕES DE OPERAÇÃO
      G1L : Bool;   // GRUPO LIGADO
      G2L : Bool;   // GRUPO LIGADO
      TEROD : Int;   // TEMPOPARA RODÍZIO DAS BOMBAS
      LIGP : Bool;   // LIGA BOMBA PRINCIPAL
      LIGC1 : Bool;   // LIGA BOMBA COMPLEMENTAR 1
      DESAB : Bool;   // DESABILITA FUNCIONAMENTO DOS GRUPOS
      T1S : Bool;   // PULSO A CADA 1 SEGUNDO
      DESAB_PART : Bool;   // DESABILITA RODIZIO POR PARTIDA
   END_VAR
   VAR_OUTPUT
      G1P : Bool;   // GRUPO 1 SELECIONADO COMO PRINCIPAL
      G2P : Bool;   // GRUPO 2 SELECIONADO COMO PRINCIPAL
      G1C1 : Bool;   // GRUPO 1 SELECIONADO COMO COMPLEMENTAR 1
      G2C1 : Bool;   // GRUPO 2 SELECIONADO COMO COMPLEMENTAR 1
      LG1 : Bool;   // LIGA GRUPO 1
      LG2 : Bool;   // LIGA GRUPO 2
   END_VAR
   VAR_IN_OUT
      TOG1P : DInt;   // TEMPO DE OPERAÇÃO GRUPO 1
      TOG2P : DInt;   // TEMPO DE OPERAÇÃO GRUPO 2
      TEOKG1 : Real;   // TEMPO OK GRUPO 1
      TEOKG2 : Real;   // TEMPO OK GRUPO 2
   END_VAR
   VAR
      GR1SELP : Bool;   // SELECIONADO COMO PRINCIPAL
      GR2SELP : Bool;   // SELECIONADO COMO PRINCIPAL
      GR1SELC1 : Bool;   // SELECIONADO COMO COMPLEMENTAR 1
      GR2SELC1 : Bool;   // SELECIONADO COMO COMPLEMENTAR 1
      PS1SG1 : Bool;   // AUXILIAR DE PULSO
      PS1SG2 : Bool;   // AUXILIAR DE PULSO
      PS1 : Bool;   // AUXILIAR DE PULSO
      PS2 : Bool;   // AUXILIAR DE PULSO
      FIMTEG1 : Bool;   // FIM DO TEMPO DE EXISTÊNCIA DO GRUPO 1
      FIMTEG2 : Bool;   // FIM DO TEMPO DE EXISTÊNCIA DO GRUPO 2
      SDESG1 : Bool;   // SOLICITAÇÃO DE DESLIGAMENTO
      SDESG2 : Bool;   // SOLICITAÇÃO DE DESLIGAMENTO
      GPL : Bool;   // GRUPO PRINCIPAL LIGADO
      GC1L : Bool;   // GRUPO COMPLEMENTAR 1 LIGADO
      SO_L : Bool;   // SOLICITAÇÃO DE PARTIDA
      SO_D : Bool;   // SOLICITAÇÃO DE DESLIGAMENTO
      RTEOPG1 : Bool;   // RESET TEMPO OK
      RTEOPG2 : Bool;   // RESET TEMPO OK
      TON1 : TON_TIME;   // TEMPORIZADOR
      TON2 : TON_TIME;   // TEMPORIZADOR
      TSDG1 : TON_TIME;   // TEMPORIZADOR
      TSDG2 : TON_TIME;   // TEMPORIZADOR
   END_VAR
   VAR_TEMP
      PRI12 : Bool;   // PRIORIDADE GRUPO 1
      TMROD : DInt;   // TEMPO DE RODIZIO
      TEROD_DI : DInt;   // TEMPO DE RODIZIO
      NGS : Int;   // NÚMERO DE GRUPOS SOLICITADOS
      NGF : Int;   // NÚMERO DE GRUPOS FUNCIONANDO
      AUX01 : Int;   // AUXILIAR UTILIZADO NA LÓGICA
      AUX02 : Int;   // AUXILIAR UTILIZADO NA LÓGICA
      AUX03 : Int;   // AUXILIAR UTILIZADO NA LÓGICA
      AUX04 : Int;   // AUXILIAR UTILIZADO NA LÓGICA
      AUX05 : Bool;   // AUXILIAR UTILIZADO NA LÓGICA
      AUX06 : Bool;   // AUXILIAR UTILIZADO NA LÓGICA
      ETT1 : Time;   // EFETIVO DO TEMPORIZADOR
      ETT2 : Time;   // EFETIVO DO TEMPORIZADOR
      ETTSDG2 : Time;   // EFETIVO DO TEMPORIZADOR
      ETTSDG1 : Time;   // EFETIVO DO TEMPORIZADOR
   END_VAR
   VAR_TEMP   // added for the SCL form of the ladder/FBD networks
      _w1 : Bool;
   END_VAR
BEGIN

REGION Network 1: CONVERSÃO DO SETPOINT DE TEMPO DE RODÍZIO